
   END_CASE;
   // ***************************************************************************************
   // Write DPL Data OF 4 WORDS to slave
   // ***************************************************************************************
   #stCONNECT_DPL_Write.ActiveEstablished := TRUE;
   #stCONNECT_DPL_Write.ConnectionType := 11;    // TCP
   #stCONNECT_DPL_Write.ID := #CONNECT_ID_2;
   #stCONNECT_DPL_Write.InterfaceId := 64;    // PROFINET Network
   #stCONNECT_DPL_Write.LocalPort := 0;
   #stCONNECT_DPL_Write.RemotePort := 502;   // 502 See TIA ONLINE HELP
   #stCONNECT_DPL_Write.RemoteAddress.ADDR[1] := #IP_OCTET_1;
   #stCONNECT_DPL_Write.RemoteAddress.ADDR[2] := #IP_OCTET_2;
   #stCONNECT_DPL_Write.RemoteAddress.ADDR[3] := #IP_OCTET_3;
   #stCONNECT_DPL_Write.RemoteAddress.ADDR[4] := #IP_OCTET_4;
   CASE #iState_Write_DPL OF
       0:  // DISCONNECT
           #MB_CLIENT_Instance_DPL_Write(REQ := FALSE,
                                         DISCONNECT := TRUE,
                                         MB_MODE := 1,
                                         MB_DATA_ADDR := 400001 + 6922,
                                         MB_DATA_LEN := 4,
                                         MB_DATA_PTR := #ReadData_DPL,
                                         CONNECT := #stCONNECT_DPL_Write);
           #iState_Write_DPL := #iState_Write_DPL + 1;
       1:  // CONNECT  
           #MB_CLIENT_Instance_DPL_Write(REQ := FALSE,
                                         DISCONNECT := FALSE,
                                         MB_MODE := 1,
                                         MB_DATA_ADDR := 400001 + 6922,
                                         MB_DATA_LEN := 4,
                                         MB_DATA_PTR := #WriteData_DPL,
                                         CONNECT := #stCONNECT_DPL_Write);
           IF #MB_CLIENT_Instance_DPL_Write.Connected AND NOT #MB_CLIENT_Instance_DPL_Write.BUSY THEN
               #woWriteDPL_ErrorID := 0;
               #iState_Write_DPL := #iState_Write_DPL + 1;
           ELSIF #MB_CLIENT_Instance_DPL_Write.ERROR THEN
               #woWriteDPL_ErrorID := #MB_CLIENT_Instance_DPL_Write.STATUS;
               #iState_Write_DPL := #iState_Write_DPL + 100;
           END_IF;
       2:  // Write Data
           FOR #Index := 0 TO 7 DO
               #WriteData_DPL[#Index] := #ILx2T_Ref.arOutputData[#Index];
           END_FOR;
           #MB_CLIENT_Instance_DPL_Write(REQ := TRUE,
                                         DISCONNECT := FALSE,
                                         MB_MODE := 1,
                                         MB_DATA_ADDR := 400001 + 6922,
                                         MB_DATA_LEN := 4,
                                         MB_DATA_PTR := #WriteData_DPL,
                                         CONNECT := #stCONNECT_DPL_Write);
           IF #MB_CLIENT_Instance_DPL_Write.DONE AND NOT #MB_CLIENT_Instance_DPL_Write.BUSY THEN
               #woWriteDPL_ErrorID := 0;
               #xErrorWriteDPL := FALSE;
           ELSIF #MB_CLIENT_Instance_DPL_Write.ERROR THEN
               #woWriteDPL_ErrorID := #MB_CLIENT_Instance_DPL_Write.STATUS;
               #iState_Write_DPL := #iState_Write_DPL + 100;
           END_IF;

       100..120:  // Error state
           #xErrorWriteDPL := TRUE;
           #diErrorCounter_DPL_Write := #diErrorCounter_DPL_Write + 1;
           #MB_CLIENT_Instance_DPL_Write(REQ := FALSE,
                                         DISCONNECT := TRUE,
                                         MB_MODE := 1,
                                         MB_DATA_ADDR := 400001 + 6922,
                                         MB_DATA_LEN := 4,
                                         MB_DATA_PTR := #WriteData_DPL,
                                         CONNECT := #stCONNECT_DPL_Write);
           #iState_Write_DPL := 0;
   END_CASE;
   // ***************************************************************************************
   // ReadParameter
   // ***************************************************************************************
   #stCONNECT_Parameter_Read.ActiveEstablished := TRUE;
   #stCONNECT_Parameter_Read.ConnectionType := 11;    // TCP
   #stCONNECT_Parameter_Read.ID := #CONNECT_ID_3;
   #stCONNECT_Parameter_Read.InterfaceId := 64;    // PROFINET Network
   #stCONNECT_Parameter_Read.LocalPort := 0;
   #stCONNECT_Parameter_Read.RemotePort := 502;   // 502 See TIA ONLINE HELP
   #stCONNECT_Parameter_Read.RemoteAddress.ADDR[1] := #IP_OCTET_1;
   #stCONNECT_Parameter_Read.RemoteAddress.ADDR[2] := #IP_OCTET_2;
   #stCONNECT_Parameter_Read.RemoteAddress.ADDR[3] := #IP_OCTET_3;
   #stCONNECT_Parameter_Read.RemoteAddress.ADDR[4] := #IP_OCTET_4;
   CASE #iState_Read_Para OF
       0:  // DISCONNECT
           #MB_CLIENT_Instance_ParaRead(REQ := FALSE,
                                        DISCONNECT := TRUE,
                                        MB_MODE := 0,
                                        MB_DATA_ADDR := 400001 + #ILx2T_Ref.udi_ModbusAddress_Read,
                                        MB_DATA_LEN := 2,
                                        MB_DATA_PTR := #ParaRead_Value,
                                        CONNECT := #stCONNECT_Parameter_Read);
           #iState_Read_Para := #iState_Read_Para + 1;

           // **********************************************************************************************************
           // ***** Reading parameters *********************************************************************************
           // **********************************************************************************************************
       1:  // CONNECT  
           #MB_CLIENT_Instance_ParaRead(REQ := FALSE,
                                        DISCONNECT := FALSE,
                                        MB_MODE := 0,
                                        MB_DATA_ADDR := 400001 + #ILx2T_Ref.udi_ModbusAddress_Read,
                                        MB_DATA_LEN := 2,
                                        MB_DATA_PTR := #ParaRead_Value,
                                        CONNECT := #stCONNECT_Parameter_Read);
           IF #MB_CLIENT_Instance_ParaRead.Connected AND NOT #MB_CLIENT_Instance_ParaRead.BUSY THEN
               #iState_Read_Para := #iState_Read_Para + 1;
           ELSIF #MB_CLIENT_Instance_ParaRead.ERROR THEN
               #woReadParameter_ErrorID := #MB_CLIENT_Instance_ParaRead.STATUS;
               #iState_Read_Para := #iState_Read_Para + 100;
           END_IF;
       2:  // Read Parameter
           IF #ILx2T_Ref.x_CommandReadParameter THEN
               #iState_Read_Para := #iState_Read_Para + 1;
           ELSE
               // #woReadParameter_ErrorID := 0;
               #xErrorReadParameter := FALSE;
           END_IF;
       3:  // Read Parameter  
           IF NOT #ILx2T_Ref.x_CommandReadParameter THEN
               #MB_CLIENT_Instance_ParaRead(REQ := FALSE,
                                            DISCONNECT := FALSE,
                                            MB_MODE := 0,
                                            MB_DATA_ADDR := 400001 + #ILx2T_Ref.udi_ModbusAddress_Read,
                                            MB_DATA_LEN := 2,
                                            MB_DATA_PTR := #ParaRead_Value,
                                            CONNECT := #stCONNECT_Parameter_Read);
               #woReadParameter_ErrorID := 0;
               #ILx2T_Ref.di_ParameterReadValue := 0;
               #ILx2T_Ref.x_StatusReadParameter_OK := FALSE;
               #iState_Read_Para := #iState_Read_Para - 1;
           ELSIF #ILx2T_Ref.x_CommandReadParameter THEN
               #MB_CLIENT_Instance_ParaRead(REQ := TRUE,
                                            DISCONNECT := FALSE,
                                            MB_MODE := 0,
                                            MB_DATA_ADDR := 400001 + #ILx2T_Ref.udi_ModbusAddress_Read,
                                            MB_DATA_LEN := 2,
                                            MB_DATA_PTR := #ParaRead_Value,
                                            CONNECT := #stCONNECT_Parameter_Read);
               IF #MB_CLIENT_Instance_ParaRead.DONE AND NOT #MB_CLIENT_Instance_ParaRead.BUSY THEN
                   #woReadParameter_ErrorID := 0;
                   #xErrorReadParameter := FALSE;
                   #ILx2T_Ref.di_ParameterReadValue := #ParaRead_Value;
                   #ILx2T_Ref.x_StatusReadParameter_OK := TRUE;
               ELSIF #MB_CLIENT_Instance_ParaRead.ERROR THEN
                   #woReadParameter_ErrorID := #MB_CLIENT_Instance_ParaRead.STATUS;
                   #ILx2T_Ref.x_StatusReadParameter_Error := TRUE;
                   #iState_Read_Para := #iState_Read_Para + 100;
               END_IF;
           END_IF;

       100..120:  // Error state
           #xErrorReadParameter := TRUE;
           #diErrorCounter_Para_Read := #diErrorCounter_Para_Read + 1;
           #MB_CLIENT_Instance_ParaRead(REQ := FALSE,
                                        DISCONNECT := TRUE,
                                        MB_MODE := 0,
                                        MB_DATA_ADDR := 400001 + #ILx2T_Ref.udi_ModbusAddress_Read,
                                        MB_DATA_LEN := 2,
                                        MB_DATA_PTR := #ParaRead_Value,
                                        CONNECT := #stCONNECT_Parameter_Read);
           #iState_Read_Para := 0;
   END_CASE;
   // ***************************************************************************************
   // WriteParameter
   // ***************************************************************************************
   #stCONNECT_Parameter_Write.ActiveEstablished := TRUE;
   #stCONNECT_Parameter_Write.ConnectionType := 11;    // TCP
   #stCONNECT_Parameter_Write.ID := #CONNECT_ID_4;
   #stCONNECT_Parameter_Write.InterfaceId := 64;    // PROFINET Network
   #stCONNECT_Parameter_Write.LocalPort := 0;
   #stCONNECT_Parameter_Write.RemotePort := 502;   // 502 See TIA ONLINE HELP
   #stCONNECT_Parameter_Write.RemoteAddress.ADDR[1] := #IP_OCTET_1;
   #stCONNECT_Parameter_Write.RemoteAddress.ADDR[2] := #IP_OCTET_2;
   #stCONNECT_Parameter_Write.RemoteAddress.ADDR[3] := #IP_OCTET_3;
   #stCONNECT_Parameter_Write.RemoteAddress.ADDR[4] := #IP_OCTET_4;
   CASE #iState_Write_Para OF
       0:  // DISCONNECT
           #MB_CLIENT_Instance_ParaWrite(REQ := FALSE,
                                         DISCONNECT := TRUE,
                                         MB_MODE := 1,
                                         MB_DATA_ADDR := 400001 + #ILx2T_Ref.udi_ModbusAddress_Write,
                                         MB_DATA_LEN := 2,
                                         MB_DATA_PTR := #ParaWrite_Value,
                                         CONNECT := #stCONNECT_Parameter_Write);
           #iState_Write_Para := #iState_Write_Para + 1;
       1:  // Write Data
           IF #ILx2T_Ref.x_CommandWriteParameter AND NOT #ILx2T_Ref.x_Status_WriteParameter_OK AND NOT #ILx2T_Ref.x_Status_WriteParameter_Error THEN
               #iState_Write_Para := 2;
           ELSE
               #xErrorWriteParameter := FALSE;
           END_IF;
           // **********************************************************************************************************
           // ***** Writing parameters *********************************************************************************
           // **********************************************************************************************************
       2:  // CONNECT  
           #ParaWrite_Value := #ILx2T_Ref.di_ParameterWriteValue;
           #MB_CLIENT_Instance_ParaWrite(REQ := FALSE,
                                         DISCONNECT := FALSE,
                                         MB_MODE := 1,
                                         MB_DATA_ADDR := 400001 + #ILx2T_Ref.udi_ModbusAddress_Write,
                                         MB_DATA_LEN := 2,
                                         MB_DATA_PTR := #ParaWrite_Value,
                                         CONNECT := #stCONNECT_Parameter_Write);
           IF #MB_CLIENT_Instance_ParaWrite.Connected AND NOT #MB_CLIENT_Instance_ParaWrite.BUSY THEN
               #woWriteParameter_ErrorID := 0;
               #iState_Write_Para := #iState_Write_Para + 1;
           ELSIF #MB_CLIENT_Instance_ParaWrite.ERROR THEN
               #woWriteParameter_ErrorID := #MB_CLIENT_Instance_ParaWrite.STATUS;
               #iState_Write_Para := #iState_Write_Para + 100;
           END_IF;
       3:  // Write Parameter
           #ParaWrite_Value := #ILx2T_Ref.di_ParameterWriteValue;
           #MB_CLIENT_Instance_ParaWrite(REQ := TRUE,
                                         DISCONNECT := FALSE,
                                         MB_MODE := 1,
                                         MB_DATA_ADDR := 400001 + #ILx2T_Ref.udi_ModbusAddress_Write,
                                         MB_DATA_LEN := 2,
                                         MB_DATA_PTR := #ParaWrite_Value,
                                         CONNECT := #stCONNECT_Parameter_Write);
           IF #MB_CLIENT_Instance_ParaWrite.DONE AND NOT #MB_CLIENT_Instance_ParaWrite.BUSY THEN
               #woWriteParameter_ErrorID := 0;
               #xErrorWriteParameter := FALSE;
               #MB_CLIENT_Instance_ParaWrite(REQ := FALSE,
                                             DISCONNECT := FALSE,
                                             MB_MODE := 1,
                                             MB_DATA_ADDR := 400001 + #ILx2T_Ref.udi_ModbusAddress_Write,
                                             MB_DATA_LEN := 2,
                                             MB_DATA_PTR := #ParaWrite_Value,
                                             CONNECT := #stCONNECT_Parameter_Write);
               #ILx2T_Ref.x_Status_WriteParameter_OK := TRUE;
               #iState_Write_Para := 1;
           ELSIF #MB_CLIENT_Instance_ParaWrite.ERROR THEN
               #ILx2T_Ref.x_Status_WriteParameter_Error := TRUE;
               #woWriteParameter_ErrorID := #MB_CLIENT_Instance_ParaWrite.STATUS;
               #iState_Write_Para := #iState_Write_Para + 100;
           END_IF;

       100..120:  // Error state
           #xErrorWriteParameter := TRUE;
           #diErrorCounter_Para_Write := #diErrorCounter_Para_Write + 1;
           #MB_CLIENT_Instance_ParaWrite(REQ := FALSE,
                                         DISCONNECT := TRUE,
                                         MB_MODE := 1,
                                         MB_DATA_ADDR := 400001 + #ILx2T_Ref.udi_ModbusAddress_Write,
                                         MB_DATA_LEN := 2,
                                         MB_DATA_PTR := #ParaWrite_Value,
                                         CONNECT := #stCONNECT_Parameter_Write);
           #iState_Write_Para := 0;

   END_CASE;

   // ********************************************************************************************
   // Communication OK or Error
   // ********************************************************************************************
   IF NOT #xErrorReadDPL AND NOT #xErrorWriteDPL AND NOT #xErrorReadParameter AND NOT #xErrorWriteParameter THEN
       #Com_OK := TRUE;
       #Error := FALSE;
   ELSE
       #Com_OK := FALSE;
       #Error := TRUE;
   END_IF;
   // ********************************************************************************************
   // Time measurements
   // Only for Diagnostic
   // ********************************************************************************************
   CASE #iStateTimeReadDPL OF
       0:
           IF #MB_CLIENT_Instance_DPL_Read.DONE THEN
               #T_ReadDPL(IN := FALSE,
                          PT := t#2m);
               #T_ReadDPL(IN := TRUE,
                          PT := t#2m);
               #iStateTimeReadDPL := #iStateTimeReadDPL + 1;
           END_IF;
       1:
           #T_ReadDPL(IN := TRUE,
                      PT := t#2m);
           IF #MB_CLIENT_Instance_DPL_Read.DONE THEN
               #t_ReadDPL_Act := #T_ReadDPL.ET;
               IF #t_ReadDPL_Act > #t_ReadDPL_Max THEN
                   #t_ReadDPL_Max := #t_ReadDPL_Act;
               ELSIF #t_ReadDPL_Act < #t_ReadDPL_Min THEN
                   #t_ReadDPL_Min := #t_ReadDPL_Act;
               END_IF;
               #T_ReadDPL(IN := FALSE,
                          PT := t#2m);
               #T_ReadDPL(IN := TRUE,
                          PT := t#2m);
           END_IF;
   END_CASE;


   CASE #iStateTimeWriteDPL OF
       0:
           IF #MB_CLIENT_Instance_DPL_Write.DONE THEN
               #T_WriteDPL(IN := FALSE,
                           PT := t#2m);
               #T_WriteDPL(IN := TRUE,
                           PT := t#2m);
               #iStateTimeWriteDPL := #iStateTimeWriteDPL + 1;
           END_IF;
       1:
           #T_WriteDPL(IN := TRUE,
                       PT := t#2m);
           IF #MB_CLIENT_Instance_DPL_Write.DONE THEN
               #t_WriteDPL_Act := #T_WriteDPL.ET;
               IF #t_WriteDPL_Act > #t_WriteDPL_Max THEN
                   #t_WriteDPL_Max := #t_WriteDPL_Act;
               ELSIF #t_WriteDPL_Act < #t_WriteDPL_Min THEN
                   #t_WriteDPL_Min := #t_WriteDPL_Act;
               END_IF;
               #T_WriteDPL(IN := FALSE,
                           PT := t#2m);
               #T_WriteDPL(IN := TRUE,
                           PT := t#2m);
           END_IF;
   END_CASE;
END_FUNCTION_BLOCK

// folder: Subroutine

FUNCTION_BLOCK "GP_OB_Initialize"   // FB2, SCL
TITLE = OB Service flags
{ S7_Optimized_Access := 'TRUE' }
AUTHOR : Cigliutt
FAMILY : GP
VERSION : 1.1
// This FB will provide the following information: 1# OB duration time 2# Timer clock and OS. IMPORTANT!!! This FB must be initialized each OB100 call, and must be called for each OB!
   VAR_INPUT
      IN_xInitialize : Bool;   // Initialize values (OB100 call)
   END_VAR
   VAR
      STC_rlLastExecValue_s : LReal;   // Last execution tick value [s]
      STC_rlReminder_s : Real;   // Reminder from last execution [ms]
      STC_dElapsed_100ms_ms : DInt;   // Elapsed time for 0.1s
      STC_dElapsed_200ms_ms : DInt;   // Elapsed time for 0.2s
      STC_dElapsed_400ms_ms : DInt;   // Elapsed time for 0.4s
      STC_dElapsed_500ms_ms : DInt;   // Elapsed time for 0.5s
      STC_dElapsed_800ms_ms : DInt;   // Elapsed time for 0.8s
      STC_dElapsed_1s_ms : DInt;   // Elapsed time for 1s
      STC_dElapsed_2s_ms : DInt;   // Elapsed time for 2s
      STC_dElapsed_5s_ms : DInt;   // Elapsed time for 5s
      STC_dElapsed_10s_ms : DInt;   // Elapsed time for 10s
      STC_dElapsed_30s_ms : DInt;   // Elapsed time for 30s
      STC_dElapsed_1min_ms : DInt;   // Elapsed time for 1min
      STC_dElapsed_2min_ms : DInt;   // Elapsed time for 2min
      STC_dElapsed_10min_ms : DInt;   // Elapsed time for 10min
      STC_dElapsed_30min_ms : DInt;   // Elapsed time for 30min
      STC_dElapsed_1h_ms : DInt;   // Elapsed time for 1h
      OUT_dExecutionTime_ms : DInt;   // OB Execution time [ms]
      OUT_dMinExecutionTime_ms : DInt;   // OB Maximum execution time [ms]
      OUT_dMaxExecutionTime_ms : DInt;   // OB Minimum execution time [ms]
      OUT_xOs_100ms : Bool;   // OS each 100ms
      OUT_xOs_200ms : Bool;   // OS each 200ms
      OUT_xOs_400ms : Bool;   // OS each 400ms
      OUT_xOs_500ms : Bool;   // OS each 500ms
      OUT_xOs_800ms : Bool;   // OS each 800ms
      OUT_xOs_1s : Bool;   // OS each 1s
      OUT_xOs_2s : Bool;   // OS each 2s
      OUT_xOs_5s : Bool;   // OS each 5s
      OUT_xOs_10s : Bool;   // OS each 10s
      OUT_xOs_30s : Bool;   // OS each 30s
      OUT_xOs_1min : Bool;   // OS each 1min
      OUT_xOs_2min : Bool;   // OS each 2min
      OUT_xOs_10min : Bool;   // OS each 10min
      OUT_xOs_30min : Bool;   // OS each 30min
      OUT_xOs_1h : Bool;   // OS each 1h
      OUT_xClock_100ms : Bool;   // Clock 100ms
      OUT_xClock_200ms : Bool;   // Clock 200ms
      OUT_xClock_400ms : Bool;   // Clock 400ms
      OUT_xClock_500ms : Bool;   // Clock 500ms
      OUT_xClock_800ms : Bool;   // Clock 800ms
      OUT_xClock_1s : Bool;   // Clock 1s
      OUT_xClock_2s : Bool;   // Clock 2s
      OUT_xClock_5s : Bool;   // Clock 5s
      OUT_xClock_10s : Bool;   // Clock 10s
      OUT_xClock_30s : Bool;   // Clock 30s
      OUT_xClock_1min : Bool;   // Clock 1min
      OUT_xClock_2min : Bool;   // Clock 2min
      OUT_xClock_10min : Bool;   // Clock 10min
      OUT_xClock_30min : Bool;   // Clock 30min
      OUT_xClock_1h : Bool;   // Clock 1h
      OUT_xDebugOFF : Bool;   // Commisioning bit - Always OFF
      OUT_xDebugON : Bool;   // Commisioning bit - Always ON
   END_VAR
   VAR_TEMP
      TMP_rlActualExecutionTime : Real;   // ActualExecutionTime [ms]
      TMP_rlActualExecutionTimeRound : Real;   // Rounded execution time [ms]
      TMP_rlActualExecutionTimeCalculated : Real;
   END_VAR
   VAR CONSTANT
      CONST_DTICK_100MS : DInt := 100;
      CONST_DTICK_200MS : DInt := 200;
      CONST_DTICK_400MS : DInt := 400;
      CONST_DTICK_500MS : DInt := 500;
      CONST_DTICK_800MS : DInt := 800;
      CONST_DTICK_1S : DInt := 1000;
      CONST_DTICK_2S : DInt := 2000;
      CONST_DTICK_5S : DInt := 5000;
      CONST_DTICK_10S : DInt := 10000;
      CONST_DTICK_30S : DInt := 30000;
      CONST_DTICK_1MIN : DInt := 60000;
      CONST_DTICK_2MIN : DInt := 120000;
      CONST_DTICK_10MIN : DInt := 600000;
      CONST_DTICK_30MIN : DInt := 1800000;
      CONST_DTICK_1H : DInt := 86400000;
      CONST_DMAX_INT : DInt := 16#7FFF_FFFF;
   END_VAR
BEGIN
   //Initialize OS bits
   #OUT_xOs_100ms := false;
   #OUT_xOs_200ms := false;
   #OUT_xOs_400ms := false;
   #OUT_xOs_500ms := false;
   #OUT_xOs_800ms := false;
   #OUT_xOs_1s := false;
   #OUT_xOs_2s := false;
   #OUT_xOs_5s := false;
   #OUT_xOs_10s := false;
   #OUT_xOs_30s := false;
   #OUT_xOs_1min := false;
   #OUT_xOs_2min := false;
   #OUT_xOs_10min := false;
   #OUT_xOs_30min := false;
   #OUT_xOs_1h := false;

   //Initialize FB execution
   IF #IN_xInitialize = true THEN


       #IN_xInitialize := false;

       #OUT_dExecutionTime_ms := 0;
       #OUT_dMinExecutionTime_ms := #CONST_DMAX_INT;
       #OUT_dMaxExecutionTime_ms := 0;
       #OUT_xClock_100ms := false;
       #OUT_xClock_200ms := false;
       #OUT_xClock_400ms := false;
       #OUT_xClock_500ms := false;
       #OUT_xClock_800ms := false;
       #OUT_xClock_1s := false;
       #OUT_xClock_2s := false;
       #OUT_xClock_5s := false;
       #OUT_xClock_10s := false;
       #OUT_xClock_30s := false;
       #OUT_xClock_1min := false;
       #OUT_xClock_2min := false;
       #OUT_xClock_10min := false;
       #OUT_xClock_30min := false;
       #OUT_xClock_1h := false;

       #STC_dElapsed_100ms_ms := 0;
       #STC_dElapsed_200ms_ms := 0;
       #STC_dElapsed_400ms_ms := 0;
       #STC_dElapsed_500ms_ms := 0;
       #STC_dElapsed_800ms_ms := 0;
       #STC_dElapsed_1s_ms := 0;
       #STC_dElapsed_2s_ms := 0;
       #STC_dElapsed_5s_ms := 0;
       #STC_dElapsed_10s_ms := 0;
       #STC_dElapsed_30s_ms := 0;
       #STC_dElapsed_1min_ms := 0;
       #STC_dElapsed_2min_ms := 0;
       #STC_dElapsed_10min_ms := 0;
       #STC_dElapsed_30min_ms := 0;
       #STC_dElapsed_1h_ms := 0;
       #STC_rlLastExecValue_s := 0;

   END_IF;
   //***** CALCULATE OB EXECUTION TIME ***** 
   //Take the execution time from the CPU
   #TMP_rlActualExecutionTime := LREAL_TO_REAL(RUNTIME(MEM := #STC_rlLastExecValue_s));

   //Convert from [s] to [ms]
   #TMP_rlActualExecutionTime := #TMP_rlActualExecutionTime * 1000.0;

   //Add the reminder of the last cycle
   #TMP_rlActualExecutionTimeCalculated := #TMP_rlActualExecutionTime + #STC_rlReminder_s;
   //Calculate the rounded value
   #TMP_rlActualExecutionTimeRound := ROUND_REAL(#TMP_rlActualExecutionTimeCalculated);
   #OUT_dExecutionTime_ms := ROUND_DINT(#TMP_rlActualExecutionTimeCalculated);

   //Save the reminder for the next cycle
   #STC_rlReminder_s := #TMP_rlActualExecutionTimeCalculated - #TMP_rlActualExecutionTimeRound;

   //Save the maximum scan value
   IF #OUT_dExecutionTime_ms > #OUT_dMaxExecutionTime_ms THEN
       #OUT_dMaxExecutionTime_ms := #OUT_dExecutionTime_ms;
   END_IF;

   //Save the minimum scan value
   IF #OUT_dExecutionTime_ms < #OUT_dMinExecutionTime_ms THEN
       #OUT_dMinExecutionTime_ms := #OUT_dExecutionTime_ms;
   END_IF;

   //***** CALCULATE SERVICES CLOCK *****

   //Increment counters for each clock
   #STC_dElapsed_100ms_ms := #STC_dElapsed_100ms_ms + #OUT_dExecutionTime_ms;
   #STC_dElapsed_200ms_ms := #STC_dElapsed_200ms_ms + #OUT_dExecutionTime_ms;
   #STC_dElapsed_400ms_ms := #STC_dElapsed_400ms_ms + #OUT_dExecutionTime_ms;
   #STC_dElapsed_500ms_ms := #STC_dElapsed_500ms_ms + #OUT_dExecutionTime_ms;
   #STC_dElapsed_800ms_ms := #STC_dElapsed_800ms_ms + #OUT_dExecutionTime_ms;
   #STC_dElapsed_1s_ms := #STC_dElapsed_1s_ms + #OUT_dExecutionTime_ms;
   #STC_dElapsed_2s_ms := #STC_dElapsed_2s_ms + #OUT_dExecutionTime_ms;
   #STC_dElapsed_5s_ms := #STC_dElapsed_5s_ms + #OUT_dExecutionTime_ms;
   #STC_dElapsed_10s_ms := #STC_dElapsed_10s_ms + #OUT_dExecutionTime_ms;
   #STC_dElapsed_30s_ms := #STC_dElapsed_30s_ms + #OUT_dExecutionTime_ms;
   #STC_dElapsed_1min_ms := #STC_dElapsed_1min_ms + #OUT_dExecutionTime_ms;
   #STC_dElapsed_2min_ms := #STC_dElapsed_2min_ms + #OUT_dExecutionTime_ms;
   #STC_dElapsed_10min_ms := #STC_dElapsed_10min_ms + #OUT_dExecutionTime_ms;
   #STC_dElapsed_30min_ms := #STC_dElapsed_30min_ms + #OUT_dExecutionTime_ms;
   #STC_dElapsed_1h_ms := #STC_dElapsed_1h_ms + #OUT_dExecutionTime_ms;

   //Calculate the 100ms
   IF #STC_dElapsed_100ms_ms >= #CONST_DTICK_100MS THEN
       #STC_dElapsed_100ms_ms := #STC_dElapsed_100ms_ms - #CONST_DTICK_100MS;

       #OUT_xOs_100ms := true;

       IF (#OUT_xClock_100ms = false) THEN
           #OUT_xClock_100ms := true;
       ELSE
           #OUT_xClock_100ms := false;
       END_IF;
   END_IF;

   //Calculate the 200ms
   IF #STC_dElapsed_200ms_ms >= #CONST_DTICK_200MS THEN
       #STC_dElapsed_200ms_ms := #STC_dElapsed_200ms_ms - #CONST_DTICK_200MS;

       #OUT_xOs_200ms := true;

       IF (#OUT_xClock_200ms = false) THEN
           #OUT_xClock_200ms := true;
       ELSE
           #OUT_xClock_200ms := false;
       END_IF;
   END_IF;

   //Calculate the 400ms
   IF #STC_dElapsed_400ms_ms >= #CONST_DTICK_400MS THEN
       #STC_dElapsed_400ms_ms := #STC_dElapsed_400ms_ms - #CONST_DTICK_400MS;

       #OUT_xOs_400ms := true;

       IF (#OUT_xClock_400ms = false) THEN
           #OUT_xClock_400ms := true;
       ELSE
           #OUT_xClock_400ms := false;
       END_IF;
   END_IF;

   //Calculate the 500ms
   IF #STC_dElapsed_500ms_ms >= #CONST_DTICK_500MS THEN
       #STC_dElapsed_500ms_ms := #STC_dElapsed_500ms_ms - #CONST_DTICK_500MS;

       #OUT_xOs_500ms := true;

       IF (#OUT_xClock_500ms = false) THEN
           #OUT_xClock_500ms := true;
       ELSE
           #OUT_xClock_500ms := false;
       END_IF;
   END_IF;

   //Calculate the 800ms
   IF #STC_dElapsed_800ms_ms >= #CONST_DTICK_800MS THEN
       #STC_dElapsed_800ms_ms := #STC_dElapsed_800ms_ms - #CONST_DTICK_800MS;

       #OUT_xOs_800ms := true;

       IF (#OUT_xClock_800ms = false) THEN
           #OUT_xClock_800ms := true;
       ELSE
           #OUT_xClock_800ms := false;
       END_IF;
   END_IF;

   //Calculate the 1s
   IF #STC_dElapsed_1s_ms >= #CONST_DTICK_1S THEN
       #STC_dElapsed_1s_ms := #STC_dElapsed_1s_ms - #CONST_DTICK_1S;

       #OUT_xOs_1s := true;

       IF (#OUT_xClock_1s = false) THEN
           #OUT_xClock_1s := true;
       ELSE
           #OUT_xClock_1s := false;
       END_IF;
   END_IF;

   //Calculate the 2s
   IF #STC_dElapsed_2s_ms >= #CONST_DTICK_2S THEN
       #STC_dElapsed_2s_ms := #STC_dElapsed_2s_ms - #CONST_DTICK_2S;

       #OUT_xOs_2s := true;

       IF (#OUT_xClock_2s = false) THEN
           #OUT_xClock_2s := true;
       ELSE
           #OUT_xClock_2s := false;
       END_IF;
   END_IF;

   //Calculate the 5s
   IF #STC_dElapsed_5s_ms >= #CONST_DTICK_5S THEN
       #STC_dElapsed_5s_ms := #STC_dElapsed_5s_ms - #CONST_DTICK_5S;

       #OUT_xOs_5s := true;

       IF (#OUT_xClock_5s = false) THEN
           #OUT_xClock_5s := true;
       ELSE
           #OUT_xClock_5s := false;
       END_IF;
   END_IF;

   //Calculate the 10s
   IF #STC_dElapsed_10s_ms >= #CONST_DTICK_10S THEN
       #STC_dElapsed_10s_ms := #STC_dElapsed_10s_ms - #CONST_DTICK_10S;

       #OUT_xOs_10s := true;

       IF (#OUT_xClock_10s = false) THEN
           #OUT_xClock_10s := true;
       ELSE
           #OUT_xClock_10s := false;
       END_IF;
   END_IF;

   //Calculate the 30s
   IF #STC_dElapsed_30s_ms >= #CONST_DTICK_30S THEN
       #STC_dElapsed_30s_ms := #STC_dElapsed_30s_ms - #CONST_DTICK_30S;

       #OUT_xOs_30s := true;

       IF (#OUT_xClock_30s = false) THEN
           #OUT_xClock_30s := true;
       ELSE
           #OUT_xClock_30s := false;
       END_IF;
   END_IF;

   //Calculate the 1min
   IF #STC_dElapsed_1min_ms >= #CONST_DTICK_1MIN THEN
       #STC_dElapsed_1min_ms := #STC_dElapsed_1min_ms - #CONST_DTICK_1MIN;

       #OUT_xOs_1min := true;

       IF (#OUT_xClock_1min = false) THEN
           #OUT_xClock_1min := true;
       ELSE
           #OUT_xClock_1min := false;
       END_IF;
   END_IF;

   //Calculate the 2min
   IF #STC_dElapsed_2min_ms >= #CONST_DTICK_2MIN THEN
       #STC_dElapsed_2min_ms := #STC_dElapsed_2min_ms - #CONST_DTICK_2MIN;

       #OUT_xOs_2min := true;

       IF (#OUT_xClock_2min = false) THEN
           #OUT_xClock_2min := true;
       ELSE
           #OUT_xClock_2min := false;
       END_IF;
   END_IF;

   //Calculate the 10min
   IF #STC_dElapsed_10min_ms >= #CONST_DTICK_10MIN THEN
       #STC_dElapsed_10min_ms := #STC_dElapsed_10min_ms - #CONST_DTICK_10MIN;

       #OUT_xOs_10min := true;

       IF (#OUT_xClock_10min = false) THEN
           #OUT_xClock_10min := true;
       ELSE
           #OUT_xClock_10min := false;
       END_IF;
   END_IF;

   //Calculate the 30min
   IF #STC_dElapsed_30min_ms >= #CONST_DTICK_30MIN THEN
       #STC_dElapsed_30min_ms := #STC_dElapsed_30min_ms - #CONST_DTICK_30MIN;

       #OUT_xOs_30min := true;

       IF (#OUT_xClock_30min = false) THEN
           #OUT_xClock_30min := true;
       ELSE
           #OUT_xClock_30min := false;
       END_IF;
   END_IF;

   //Calculate the 1h
   IF #STC_dElapsed_1h_ms >= #CONST_DTICK_1H THEN
       #STC_dElapsed_1h_ms := #STC_dElapsed_1h_ms - #CONST_DTICK_1H;

       #OUT_xOs_1h := true;

       IF (#OUT_xClock_1h = false) THEN
           #OUT_xClock_1h := true;
       ELSE
           #OUT_xClock_1h := false;
       END_IF;
   END_IF;
END_FUNCTION_BLOCK

FUNCTION "GP_GetArraySize" : Int   // FC9, SCL
{ S7_Optimized_Access := 'TRUE' }
AUTHOR : Cigliutt
FAMILY : GP
VERSION : 1.0
   VAR_IN_OUT
      INO_vArray : Variant;
   END_VAR
   VAR_TEMP
      TMP_udNumEl : UDInt;
   END_VAR
BEGIN
   #TMP_udNumEl := 0;

   IF IS_ARRAY(#INO_vArray) THEN
       #TMP_udNumEl := CountOfElements(#INO_vArray);
   END_IF;

   #GP_GetArraySize := UDINT_TO_INT(#TMP_udNumEl);
END_FUNCTION

FUNCTION "GP_BlockMoveStruct" : Int   // FC13, SCL
{ S7_Optimized_Access := 'TRUE' }
AUTHOR : Cigliutt
FAMILY : GP
VERSION : 1.0
   VAR_INPUT
      IN_iSourceIndex : Int;
      IN_iDestIndex : Int;
      IN_iCount : Int;
   END_VAR
   VAR_IN_OUT
      INO_vSourceArrayStruct : Variant;
      INO_vDestArrayStruct : Variant;
   END_VAR
BEGIN
   #GP_BlockMoveStruct :=  MOVE_BLK_VARIANT(SRC:=#INO_vSourceArrayStruct,
                                            COUNT:=INT_TO_UDINT(#IN_iCount),
                                            SRC_INDEX:=INT_TO_DINT(#IN_iSourceIndex),
                                            DEST_INDEX:=INT_TO_DINT(#IN_iDestIndex),
                                            DEST=>#INO_vDestArrayStruct);
END_FUNCTION

// folder: TaskErrors

ORGANIZATION_BLOCK "Time error interrupt"   // OB80, LAD, TimeErrorInterrupt
{ S7_Optimized_Access := 'TRUE' }
VERSION : 0.1
   VAR_INPUT
      Fault_ID : Byte;   // Fault identifier
      Csg_OBnr : OB_Any;   // Number of OB causing the error
      Csg_Prio : UInt;   // Priority of OB causing the error
   END_VAR
BEGIN
END_ORGANIZATION_BLOCK

ORGANIZATION_BLOCK "Diagnostic error interrupt"   // OB82, LAD, DiagnosticErrorInterrupt
{ S7_Optimized_Access := 'TRUE' }
VERSION : 0.1
   VAR_INPUT
      IO_State : Word;   // IO state of the HW object
      LADDR : Hw_Any;   // Hardware identifier
      Channel : UInt;   // Channel number
      MultiError : Bool;   // =true if more than one error is present
   END_VAR
   VAR_TEMP
      RALM : Struct
         AINFO : "AINFO_";
         TINFO : "TINFO_";
         RETVAL : Int;
         ALLARMI_da_OB82 : Struct
            RALM : "PN_Alarm";
            LADDR : Hw_Any;
            evento_uscente : Bool;
         END_STRUCT;
      END_STRUCT;
      TMP_dId : DInt;
   END_VAR
BEGIN

REGION Network 1
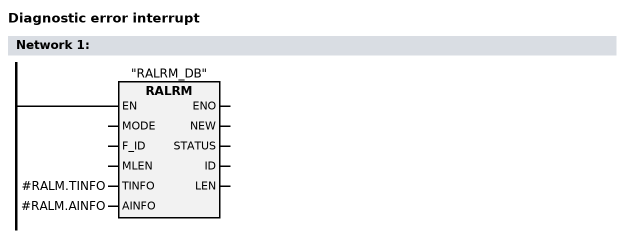
   "RALRM_DB"(TINFO := #RALM.TINFO, AINFO := #RALM.AINFO);   // RALRM
END_REGION

REGION Network 2 (SCL): Set alarms
   #TMP_dId:=UINT_TO_DINT("RALRM_DB".ID);

   IF "RALRM_DB".NEW THEN
       CASE #TMP_dId OF
           1:
               "RALRM_AUX_DB".tAlm.tF.xDevice1 := 1;
           2:
               "RALRM_AUX_DB".tAlm.tF.xDevice2 := 1;
           3:
               "RALRM_AUX_DB".tAlm.tF.xDevice3 := 1;
           4:
               "RALRM_AUX_DB".tAlm.tF.xDevice4 := 1;
           5:
               "RALRM_AUX_DB".tAlm.tF.xDevice5 := 1;
           6:
               "RALRM_AUX_DB".tAlm.tF.xDevice6 := 1;
           7:
               "RALRM_AUX_DB".tAlm.tF.xDevice7 := 1;
           8:
               "RALRM_AUX_DB".tAlm.tF.xDevice8 := 1;
           9:
               "RALRM_AUX_DB".tAlm.tF.xDevice9 := 1;
           10:
               "RALRM_AUX_DB".tAlm.tF.xDevice10 := 1;
           ELSE
               ;
       END_CASE;
   END_IF;
END_REGION
END_ORGANIZATION_BLOCK

ORGANIZATION_BLOCK "Pull or plug of modules"   // OB83, LAD, PullPlug
{ S7_Optimized_Access := 'TRUE' }
VERSION : 0.1
   VAR_INPUT
      LADDR : Hw_Io;   // Hardware identifier
      Event_Class : Byte;   // 16#38/39: module inserted, removed
      Fault_ID : Byte;   // Fault identifier
   END_VAR
BEGIN
END_ORGANIZATION_BLOCK

ORGANIZATION_BLOCK "Rack or station failure"   // OB86, LAD, RackStationFailure
{ S7_Optimized_Access := 'TRUE' }
VERSION : 0.1
   VAR_INPUT
      LADDR : Hw_Device;   // Hardware identifier
      Event_Class : Byte;   // Event class
      Fault_ID : Byte;   // Fault identifier
   END_VAR
BEGIN
END_ORGANIZATION_BLOCK

ORGANIZATION_BLOCK "Programming error"   // OB121, LAD, ProgrammingError
{ S7_Optimized_Access := 'TRUE' }
VERSION : 0.1
   VAR_INPUT
      BlockNr : UInt;   // Number of causing block
      Reaction : USInt;   // 0:ignore, 1:substitute, 2:skip
      Fault_ID : Byte;   // Fault identifier
      BlockType : USInt;   // 16#01:OB, 16#02:FC, 16#03:FB, 16#04:SFC, 16#05:SFB, 16#06:DB: Type of block causing the error
      Area : USInt;   // Area where the error occured
      DBNr : DB_ANY;   // DB number if Area = DB or DI
      Csg_OBNr : OB_Any;   // Number of OB causing the error
      Csg_Prio : USInt;   // Priority of OB causing the error
      Width : USInt;   // 0:bit, 1:byte, 2:word, 3:dword, 4:lword
   END_VAR
BEGIN
END_ORGANIZATION_BLOCK

ORGANIZATION_BLOCK "IO access error"   // OB122, LAD, IOAccessError
{ S7_Optimized_Access := 'TRUE' }
VERSION : 0.1
   VAR_INPUT
      BlockNr : UInt;   // Number of causing block
      Reaction : USInt;   // 0:ignore, 1:substitute, 2:skip
      Fault_ID : Byte;   // 16#42:reading, 16#43:writing
      BlockType : USInt;   // 16#01:OB, 16#02:FC, 16#03:FB, 16#04:SFC, 16#05:SFB, 16#06:DB: Type of block causing the error
      Area : USInt;   // 16#81:I, 16#82:Q: IO area where the IOaccess error occured
      DBNr : DB_ANY;   // Reserved for system
      Csg_OBNr : OB_Any;   // Number of OB causing the error
      Csg_Prio : USInt;   // Priority of OB causing the error
      Width : USInt;   // 0:bit, 1:byte, 2:word, 3:dword, 4:lword
   END_VAR
BEGIN
END_ORGANIZATION_BLOCK